screen "106_Rocno_postaja6" 1280x800, template "100_Rocno"
   IOField "I/O field_1" at 1132,158 size 125x32; FormatPattern 99999; Unit  l/min
      ProcessValue <- "FB_IOL_IFM_SV_DB_uPretok"
   IOField "I/O field_2" at 1132,210 size 128x32; FormatPattern 99.9; Unit  °C
      ProcessValue <- "FB_IOL_IFM_SV_DB_fTemperatura"
   TextField "Text field_2" at 1090,159 size 19x25; Text 'Q'
   TextField "Text field_3" at 1093,216 size 16x25; Text 'T'
   TextField "Text field_4" at 1144,120 size 58x25; Text 'VODA'
   IOField "I/O field_3" at 1132,304 size 125x32; FormatPattern 99.9; Unit  bar
      ProcessValue <- "FB_Lin_FESTO_PNEVMATIKA_PRITISK_Q_izhod"
   TextField "Text field_5" at 1090,305 size 17x25; Text 'P'
   TextField "Text field_7" at 1144,266 size 56x25; Text 'ZRAK'
   IOField "I/O field_4" at 1133,400 size 125x32; FormatPattern 99.9; Unit  bar
      ProcessValue <- "FB_FESTO_VPPM_DB_setstatZeljeniPritisk"
   TextField "Text field_6" at 1091,401 size 17x25; Text 'P'
   TextField "Text field_8" at 1100,360 size 169x25; Text 'P ZATISKOVANJA'
   TextField "Text field_17" at 613,544 size 239x46; Text 'POBIRANJE/NALAGANJE KOMADA'
   IOField "I/O field_7" at 742,605 size 133x35; FormatPattern 99.9; Unit  mm
      ProcessValue <- "DB_HMI_SDAT1_PozPobiranje"
   IOField "I/O field_8" at 739,666 size 136x35; FormatPattern 99.9; Unit  mm
      ProcessValue <- "DB_HMI_SDAT1_PozNalaganje"
   TextField "Text field_12" at 280,615 size 118x25; Text 'NALAGANJE'
   TextField "Text field_13" at 281,677 size 114x25; Text 'POBIRANJE'
   TextField "Text field_14" at 290,544 size 239x46; Text 'POBIRANJE/NALAGANJE PLOŠČICE'
   Circle "Circle_8" at 393,678 size 21x21
      Appearance <- "SDAT2_oPoz1Dosezena"
   Circle "Circle_7" at 394,618 size 21x21
      Appearance <- "SDAT2_oPoz2Dosezena"
   IOField "I/O field_10" at 421,670 size 136x32; FormatPattern 99.9; Unit  mm
      ProcessValue <- "DB_HMI_SDAT2_PozPobiranje"
   IOField "I/O field_9" at 425,613 size 133x32; FormatPattern 99.9; Unit  mm
      ProcessValue <- "DB_HMI_SDAT2_PozNalaganje"
   IOField "I/O field_12" at 422,709 size 136x32; FormatPattern 99.99; Unit  mm
      ProcessValue <- "SDAT2_out"
   TextField "Text field_11" at 434,112 size 84x25; Text 'Keyence'
   IOField "I/O field_13" at 432,190 size 109x32; FormatPattern 999999; Unit  mm
      ProcessValue <- "DB_KEYENCE_Elektroda_ZeljenaPozicija_POZ1"
   IOField "I/O field_14" at 432,244 size 109x32; FormatPattern 999999; Unit  mm
      ProcessValue <- "DB_KEYENCE_Elektroda_ZeljenaPozicija_POZ2"
   TextField "Text field_18" at 369,147 size 213x25; Text 'ELEKTRODA GOR/DOL'
   IOField "I/O field_17" at 432,290 size 109x32; FormatPattern 999999; Unit  mm
      ProcessValue <- "DB_KEYENCE_Elektroda_ZeljenaPozicija_POZ3_elektrodaStisnjena"
   IOField "I/O field_18" at 431,334 size 109x32; FormatPattern 999999; Unit  mm
      ProcessValue <- "DB_KEYENCE_Elektroda_ZeljenaPozicija_POZ4_elektrodaZavarjeno"
   TextField "Text field_9" at 282,194 size 81x25; Text 'ZGORAJ'
   TextField "Text field_19" at 282,339 size 117x25; Text 'ZAVARJENO'
   TextField "Text field_20" at 282,294 size 112x25; Text 'STISNJENO'
   TextField "Text field_21" at 282,248 size 99x25; Text 'HLAJENJE'
   Circle "Circle_1" at 398,195 size 20x20
      Appearance <- "FB_KEYENCE_GT2_ODMIKVARJENJA_oPoz1Dosezena"
   Circle "Circle_2" at 399,250 size 20x20
      Appearance <- "FB_KEYENCE_GT2_ODMIKVARJENJA_oPoz2Dosezena"
   Circle "Circle_3" at 401,296 size 20x20
      Appearance <- "FB_KEYENCE_GT2_ODMIKVARJENJA_oPoz3Dosezena"
   Circle "Circle_4" at 401,339 size 20x20
      Appearance <- "FB_KEYENCE_GT2_ODMIKVARJENJA_oPoz4Dosezena"
   IOField "I/O field_11" at 740,706 size 136x35; FormatPattern 99.99; Unit  mm
      ProcessValue <- "SDAT1_out"
   IOField "I/O field_6" at 531,408 size 128x32; FormatPattern 999999; Unit  mm
      ProcessValue <- "Keyence_OdmičniCilinderVarjenja"
   TextField "Text field_1" at 608,610 size 118x25; Text 'NALAGANJE'
   TextField "Text field_10" at 608,672 size 114x25; Text 'POBIRANJE'
   Circle "Circle_9" at 716,674 size 21x21
      Appearance <- "SDAT1_oPoz1Dosezena"
   Circle "Circle_10" at 719,612 size 21x21
      Appearance <- "SDAT1_oPoz2Dosezena"
   TextField "Text field_22" at 823,111 size 84x25; Text 'Keyence'
   TextField "Text field_23" at 691,147 size 268x25; Text 'ELEKTRODA NAZAJ/NAPREJ'
   TextField "Text field_24" at 687,194 size 67x25; Text 'NAZAJ'
   TextField "Text field_27" at 687,243 size 78x25; Text 'NAPREJ'
   IOField "I/O field_15" at 805,190 size 109x32; FormatPattern 999999; Unit  mm
      ProcessValue <- "DB_KEYENCE_Kroznik_ZeljenaPozicija_POZ1"
   IOField "I/O field_16" at 805,242 size 109x32; FormatPattern 999999; Unit  mm
      ProcessValue <- "DB_KEYENCE_Kroznik_ZeljenaPozicija_POZ2"
   IOField "I/O field_5" at 944,408 size 125x32; FormatPattern s999999; Unit  mm
      ProcessValue <- "Keyence_OdmičniCilinderKonusa"
   Circle "Circle_5" at 770,198 size 20x20
      Appearance <- "FB_KEYENCE_GT2_odmikKonusaKroznika_oPoz1Dosezena"
   Circle "Circle_6" at 770,245 size 20x20
      Appearance <- "FB_KEYENCE_GT2_odmikKonusaKroznika_oPoz2Dosezena"
   IOField "I/O field_19" at 564,190 size 105x32; FormatPattern 999999; Unit  mm
      ProcessValue <- "DB_KEYENCE_Elektroda_TOLERANCA{1}"
   IOField "I/O field_20" at 565,244 size 105x32; FormatPattern 999999; Unit  mm
      ProcessValue <- "DB_KEYENCE_Elektroda_TOLERANCA{2}"
   IOField "I/O field_21" at 564,290 size 105x32; FormatPattern 999999; Unit  mm
      ProcessValue <- "DB_KEYENCE_Elektroda_TOLERANCA{3}"
   IOField "I/O field_22" at 565,334 size 105x32; FormatPattern 999999; Unit  mm
      ProcessValue <- "DB_KEYENCE_Elektroda_TOLERANCA{4}"
   IOField "I/O field_23" at 954,190 size 106x32; FormatPattern 999999; Unit  mm
      ProcessValue <- "DB_KEYENCE_TOLERANCA{1}"
   IOField "I/O field_24" at 954,242 size 106x32; FormatPattern 999999; Unit  mm
      ProcessValue <- "DB_KEYENCE_TOLERANCA{2}"
   TextField "Text field_15" at 934,191 size 20x25; Text '+'
   TextField "Text field_16" at 937,205 size 13x25; Text '-'
   TextField "Text field_25" at 937,241 size 20x25; Text '+'
   TextField "Text field_26" at 940,255 size 13x25; Text '-'
   TextField "Text field_28" at 548,188 size 20x25; Text '+'
   TextField "Text field_29" at 551,202 size 13x25; Text '-'
   TextField "Text field_30" at 548,242 size 20x25; Text '+'
   TextField "Text field_31" at 551,256 size 13x25; Text '-'
   TextField "Text field_32" at 548,289 size 20x25; Text '+'
   TextField "Text field_33" at 551,303 size 13x25; Text '-'
   TextField "Text field_34" at 548,334 size 20x25; Text '+'
   TextField "Text field_35" at 551,348 size 13x25; Text '-'
   IOField "I/O field_25" at 1090,512 size 174x32; FormatPattern 99999; Unit  kos
      ProcessValue <- "DB_HMI_ČiščenjeElektrode_ZeljenoStevilo"
   TextField "Text field_36" at 1125,460 size 114x46; Text 'CISCENJE ELEKTRODE'

screen "41_Settings2" 1280x800, template "02_Settings"
   GraphicView "Graphic view_2" at 0,0 size 1280x800; Picture "PopUpBackground"
      Visibility <- "PopUpBackground"
   IOField "I/O field_1" at 1132,158 size 125x32; FormatPattern 99999; Unit  l/min
      ProcessValue <- "FB_IOL_IFM_SV_DB_uPretok"
   IOField "I/O field_2" at 1132,210 size 128x32; FormatPattern 99.9; Unit  °C
      ProcessValue <- "FB_IOL_IFM_SV_DB_fTemperatura"
   TextField "Text field_2" at 1090,159 size 19x25; Text 'Q'
   TextField "Text field_3" at 1093,216 size 16x25; Text 'T'
   TextField "Text field_4" at 1144,120 size 58x25; Text 'VODA'
   IOField "I/O field_3" at 1132,314 size 125x32; FormatPattern 99.9; Unit  bar
      ProcessValue <- "FB_Lin_FESTO_PNEVMATIKA_PRITISK_Q_izhod"
   TextField "Text field_5" at 1090,315 size 17x25; Text 'P'
   TextField "Text field_7" at 1144,276 size 56x25; Text 'ZRAK'
   IOField "I/O field_4" at 1132,470 size 125x32; FormatPattern 99.9; Unit  bar
      ProcessValue <- "FB_FESTO_VPPM_DB_setstatZeljeniPritisk"
   TextField "Text field_6" at 1090,471 size 17x25; Text 'P'
   TextField "Text field_8" at 1099,430 size 169x25; Text 'P ZATISKOVANJA'
   TextField "Text field_17" at 613,544 size 239x46; Text 'POBIRANJE/NALAGANJE KOMADA'
   Group "Group_2" at 606,112 size 282x342
   IOField "I/O field_7" at 742,605 size 133x35; FormatPattern 99.9; Unit  mm
      ProcessValue <- "DB_HMI_SDAT1_PozPobiranje"
   IOField "I/O field_8" at 739,666 size 136x35; FormatPattern 99.9; Unit  mm
      ProcessValue <- "DB_HMI_SDAT1_PozNalaganje"
   TextField "Text field_12" at 280,615 size 118x25; Text 'NALAGANJE'
   TextField "Text field_13" at 281,677 size 114x25; Text 'POBIRANJE'
   TextField "Text field_14" at 290,544 size 239x46; Text 'POBIRANJE/NALAGANJE PLOŠČICE'
   Circle "Circle_8" at 393,678 size 21x21
      Appearance <- "SDAT2_oPoz1Dosezena"
   Circle "Circle_7" at 394,618 size 21x21
      Appearance <- "SDAT2_oPoz2Dosezena"
   IOField "I/O field_10" at 421,670 size 136x32; FormatPattern 99.9; Unit  mm
      ProcessValue <- "DB_HMI_SDAT2_PozPobiranje"
   IOField "I/O field_9" at 425,613 size 133x32; FormatPattern 99.9; Unit  mm
      ProcessValue <- "DB_HMI_SDAT2_PozNalaganje"
   IOField "I/O field_12" at 422,709 size 136x32; FormatPattern 99.99; Unit  mm
      ProcessValue <- "SDAT2_out"
   TextField "Text field_11" at 387,114 size 84x25; Text 'Keyence'
   IOField "I/O field_13" at 432,190 size 125x32; FormatPattern 999999; Unit  um
      ProcessValue <- "DB_KEYENCE_Elektroda_ZeljenaPozicija_POZ1"
   IOField "I/O field_14" at 432,244 size 125x32; FormatPattern 999999; Unit  um
      ProcessValue <- "DB_KEYENCE_Elektroda_ZeljenaPozicija_POZ2"
   TextField "Text field_18" at 333,147 size 213x25; Text 'ELEKTRODA GOR/DOL'
   IOField "I/O field_17" at 432,290 size 125x32; FormatPattern 999999; Unit  um
      ProcessValue <- "DB_KEYENCE_Elektroda_ZeljenaPozicija_POZ3_elektrodaStisnjena"
   IOField "I/O field_18" at 431,334 size 125x32; FormatPattern 999999; Unit  um
      ProcessValue <- "DB_KEYENCE_Elektroda_ZeljenaPozicija_POZ4_elektrodaZavarjeno"
   TextField "Text field_9" at 318,194 size 81x25; Text 'ZGORAJ'
   TextField "Text field_19" at 282,339 size 117x25; Text 'ZAVARJENO'
   TextField "Text field_20" at 287,294 size 112x25; Text 'STISNJENO'
   TextField "Text field_21" at 300,248 size 99x25; Text 'HLAJENJE'
   Circle "Circle_1" at 398,195 size 20x20
      Appearance <- "FB_KEYENCE_GT2_ODMIKVARJENJA_oPoz1Dosezena"
   Circle "Circle_2" at 399,250 size 20x20
      Appearance <- "FB_KEYENCE_GT2_ODMIKVARJENJA_oPoz2Dosezena"
   Circle "Circle_3" at 401,296 size 20x20
      Appearance <- "FB_KEYENCE_GT2_ODMIKVARJENJA_oPoz3Dosezena"
   Circle "Circle_4" at 401,339 size 20x20
      Appearance <- "FB_KEYENCE_GT2_ODMIKVARJENJA_oPoz4Dosezena"
   IOField "I/O field_11" at 740,706 size 136x35; FormatPattern 99.99; Unit  mm
      ProcessValue <- "SDAT1_out"
   IOField "I/O field_6" at 428,406 size 128x32; FormatPattern s999999; Unit  um
      ProcessValue <- "Keyence_OdmičniCilinderVarjenja"
   TextField "Text field_1" at 608,610 size 118x25; Text 'NALAGANJE'
   TextField "Text field_10" at 608,672 size 114x25; Text 'POBIRANJE'
   Circle "Circle_9" at 716,674 size 21x21
      Appearance <- "SDAT1_oPoz1Dosezena"
   Circle "Circle_10" at 719,612 size 21x21
      Appearance <- "SDAT1_oPoz2Dosezena"
   TextField "Text field_22" at 703,114 size 84x25; Text 'Keyence'
   TextField "Text field_23" at 620,147 size 268x25; Text 'ELEKTRODA NAZAJ/NAPREJ'
   TextField "Text field_24" at 640,194 size 67x25; Text 'NAZAJ'
   TextField "Text field_27" at 635,243 size 78x25; Text 'NAPREJ'
   IOField "I/O field_15" at 748,190 size 125x32; FormatPattern 999999; Unit  um
      ProcessValue <- "DB_KEYENCE_Kroznik_ZeljenaPozicija_POZ1"
   IOField "I/O field_16" at 748,242 size 125x32; FormatPattern 999999; Unit  um
      ProcessValue <- "DB_KEYENCE_Kroznik_ZeljenaPozicija_POZ2"
   IOField "I/O field_5" at 748,405 size 125x32; FormatPattern s999999; Unit  um
      ProcessValue <- "Keyence_OdmičniCilinderKonusa"
   Circle "Circle_5" at 713,198 size 20x20
      Appearance <- "FB_KEYENCE_GT2_odmikKonusaKroznika_oPoz1Dosezena"
   Circle "Circle_6" at 713,245 size 20x20
      Appearance <- "FB_KEYENCE_GT2_odmikKonusaKroznika_oPoz2Dosezena"

PopupScreen "VARILNIK" 300x695
   Button "Button_1" at 48,52 size 188x72; TextOff 'RESET'
      on Release: ResetBit("DB_HMI_Varjenje_ResetWithWC")
      on Press: SetBit("DB_HMI_Varjenje_ResetWithWC")
   Button "Button_2" at 48,140 size 188x72; TextOff 'RESET + ZVAR'
   SymbolicIOField "Symbolic I/O field_1" at 43,271 size 201x29; TextOn '1'; TextOff '0'; TextList "BOSH"
      ProcessValue <- "StatusCode"
   TextField "Text field_1" at 51,99 size 176x23; Text 'Reset varilnika z WC'
   TextField "Text field_2" at 52,187 size 176x23; Text 'Reset varilnika z zvarom'
   TextField "Text field_3" at 43,244 size 176x23; Text 'STATUS VARILNIKA:'
   TextField "Text field_4" at 37,10 size 221x23; Text 'VARILNIK BOSH 6000'

PopupScreen "STEVCI" 810x660
   TextField "Text field_14" at 12,94 size 150x23; Text 'ŠTEVEC SKUPAJ'
   IOField "I/O field_5" at 193,93 size 133x32; FormatPattern 999999; Unit  KOS
      ProcessValue <- "DB_STEVCI_STEVCI_SKUPAJ"
   TextField "Text field_1" at 12,143 size 129x21; Text 'ZAVARJENO OK'
   TextField "Text field_2" at 12,182 size 141x21; Text 'ZAVARJENO NOK'
   IOField "I/O field_1" at 196,137 size 133x32; FormatPattern 999999; Unit  KOS
      ProcessValue <- "DB_STEVCI_STEVCI_ZavarjenoOK"
   IOField "I/O field_2" at 196,176 size 133x32; FormatPattern 999999; Unit  KOS
      ProcessValue <- "DB_STEVCI_STEVCI_ZavarjenoNOK"
   TextField "Text field_3" at 243,10 size 214x31; Text 'ŠTEVCI IZDELKOV'
   TextField "Text field_4" at 14,55 size 96x23; Text 'VARJENJE'
   TextField "Text field_5" at 404,94 size 150x23; Text 'ŠTEVEC SKUPAJ'
   IOField "I/O field_3" at 585,93 size 133x32; FormatPattern 999999; Unit  KOS
      ProcessValue <- "DB_STEVCI_STEVCI KAMERA_SKUPAJ"
   TextField "Text field_6" at 404,143 size 100x21; Text 'KAMERA OK'
   TextField "Text field_7" at 404,182 size 112x21; Text 'KAMERA NOK'
   IOField "I/O field_4" at 588,137 size 133x32; FormatPattern 999999; Unit  KOS
      ProcessValue <- "DB_STEVCI_STEVCI KAMERA_KameraOK"
   IOField "I/O field_6" at 588,176 size 133x32; FormatPattern 999999; Unit  KOS
      ProcessValue <- "DB_STEVCI_STEVCI KAMERA_KameraNOK"
   TextField "Text field_8" at 406,55 size 82x23; Text 'KAMERA'
   TextField "Text field_9" at 765,14 size 23x24; Text 'X'
   Button "btnPreviousScreen" at 744,0 size 66x55; TextOff 'Text'
      on Click: function_efd93a16("STEVCI", 0, 0, 0, -1, 1)

PopupScreen "RESETSKATEL" 300x695
   Button "Button_1_1" at 48,70 size 188x72; TextOff 'IZPRAZNI SKATLO 1'
      on Press: SetBit("DB_HMI_TekočiTrak_btnResetSkatle1")
      on Release: ResetBit("DB_HMI_TekočiTrak_btnResetSkatle1")
   Button "Button_2" at 43,279 size 188x72; TextOff 'IZPRAZNI SKATLO 2'
      on Press: SetBit("DB_HMI_TekočiTrak_btnResetSKatle2")
      on Release: ResetBit("DB_HMI_TekočiTrak_btnResetSKatle2")
   TextField "Text field_1" at 49,119 size 186x23; Text 'Reset stevca polne škatle'
   TextField "Text field_2" at 47,328 size 176x23; Text 'Reset števca polne škatle'
   TextField "Text field_3" at 16,154 size 176x23; Text 'STATUS :'
   TextField "Text field_4" at 10,10 size 281x23; Text 'SKATLA IZDELKOV POLNA'
   TextField "Text field_5" at 16,367 size 176x23; Text 'STATUS :'
   SymbolicIOField "Symbolic I/O field_1" at 79,155 size 191x22; TextOff '0'; TextOn '1'; TextList "StatusSkatel"
      ProcessValue <- "FB_TekociTrak_DB_stat_skatla1Polna"
   SymbolicIOField "Symbolic I/O field_2" at 79,368 size 191x22; TextOn '1'; TextOff '0'; TextList "StatusSkatel"
      ProcessValue <- "FB_TekociTrak_DB_stat_skatla2Polna"

VB script "ActivateAlarmControlScreen"
   bec8f1e5-2ab1-45f6-ad91-1d37c469eb91 20_Messages,0

VB script "ActivateStartScreen"
   HmiRuntime.BaseScreenName = SmartTags("StartScreenName")

VB script "CheckCurrentLanguage"
   If HmiRuntime.Language = 1031 Then 'German
   	SmartTags("CurrentLanguage") = 0
   	ElseIf HmiRuntime.Language = 1033 Then 'English US
   	SmartTags("CurrentLanguage") = 1
   End If
   
   	

VB script "CheckCurrentUserName"
   If SmartTags("CurrentUserName") = "" Or SmartTags("CurrentUserName") = "User Name" Or SmartTags("CurrentUserName") = "Benutzer" Then
     
     If HmiRuntime.Language = 1031 Then 'Germany
       SmartTags("CurrentUserName") = "Benutzer"
       
     ElseIf HmiRuntime.Language = 1033 Then 'English US
       SmartTags("CurrentUserName") = "User Name"
     End If
     
     SmartTags("UserIsLoggedIn") = False
   Else
     If SmartTags("CurrentUserName") <> "User Name" And SmartTags("CurrentUserName") <> "Benutzer" Then
       SmartTags("UserIsLoggedIn") = True  
     End If
   End If

VB script "CheckDiagState"
   If SmartTags("@DiagnosticsIndicatorTag") = 1 Then
   	SmartTags("DiagState") = 1
   Else
   	SmartTags("DiagState") = 0
   End If

VB script "GetStartScreenName"
   SmartTags("StartScreenName") = HmiRuntime.BaseScreenName

VB script "ShowLoginPopUp"
   efd93a16-2665-4b85-bcb9-25eddcb7b6f4 Template_Logon_Logoff,480,110,$3$hmiOn$,$3$hmiAnimationOff$,$3$hmiFast$

VB script "ShowOperatingModePopUp"
   efd93a16-2665-4b85-bcb9-25eddcb7b6f4 Template_Operating_Mode,428,110,$3$hmiOn$,$3$hmiAnimationOff$,$3$hmiFast$

VB script "ShowOptionPanelPopUp"
   efd93a16-2665-4b85-bcb9-25eddcb7b6f4 OptionPanel_4_Buttons, 890, 110, $3$hmiOn$, $3$hmiRight$, $3$hmiFast$

VB script "ShowRecipePopUp"
   efd93a16-2665-4b85-bcb9-25eddcb7b6f4 Template_Recipe,290,110,$3$hmiOn$,$3$hmiAnimationOff$,$3$hmiFast$

VB script "VBFunction_1"
   'Tip:
   ' 1. Use the <CTRL+SPACE> or <CTRL+I> shortcut to open a list of all objects and functions
   ' 2. Write the code using the HMI Runtime object.
   '  Example: HmiRuntime.Screens("Screen_1").
   ' 3. Use the <CTRL+J> shortcut to create an object reference.
   'Write the code as of this position:
   
   'Please replace all sequences which are enclosed with '_' by your own code.
   
   
   '1s trigger
   
   'Poglej ce je napaka Varjenja in prigaži meni
   
   'Rectangle_17
   
   'Dim btnResetSkatle1, btnResetSkatle2
   'Set btnResetSkatle1 = HmiRuntime.ActiveScreen.ScreenItems("Button_2")
   'Set btnResetSkatle2 = HmiRuntime.ActiveScreen.ScreenItems("Rectangle_17")
   'Set btnResetSkatle1 = HmiRuntime.Screens("Slide-in screen left").ScreenItems("Button_1")
   Dim activatescreen11
   Dim screenname,txt
   screenname = HmiRuntime.BaseScreenName
   
   'Set txt = HmiRuntime.ActiveScreen.ScreenItems("Text15")
   'txt.Text = screenname
   
   If  SmartTags("TimerReady") = 0  Then
   	'ShowSlideInScreen "Slide-in screen left", hmiOn
   	efd93a16-2665-4b85-bcb9-25eddcb7b6f4 VARILNIK,0,105,$3$hmiOn$,$3$hmiAnimationOff$,$3$hmiFast$
   	activatescreen11 = True
   	
   	
   Else
   	efd93a16-2665-4b85-bcb9-25eddcb7b6f4 VARILNIK,0,105,$3$hmiOff$,$3$hmiAnimationOff$,$3$hmiFast$
   	activatescreen11 = False
   End If
   
   
   
   'Please replace all sequences which are enclosed with '_' by your own code.
   If ((SmartTags("DB_STEVCI_STEVEC_SKATEL_SKATLA1") >= SmartTags("DB_STEVCI_STEVCI_ZELENAPOLNA_SKATLA_SKATLA1") Or (SmartTags("DB_STEVCI_STEVEC_SKATEL_SKATLA2") >= SmartTags("DB_STEVCI_STEVCI_ZELENAPOLNA_SKATLA_SKATLA2"))) And (Not activatescreen11)) Then
   	efd93a16-2665-4b85-bcb9-25eddcb7b6f4 RESETSKATEL,0,105,$3$hmiOn$,$3$hmiAnimationOff$,$3$hmiFast$
   	'btnResetSkatle1.Top = 10
   	'btnResetSkatle1.Visible = 1
   	'ModraSkatla
   	'btnResetSkatle2.BackColor = RGB(0,95,135)
   	
   	
   Else
   	efd93a16-2665-4b85-bcb9-25eddcb7b6f4 RESETSKATEL,0,105,$3$hmiOff$,$3$hmiAnimationOff$,$3$hmiFast$
   	'btnResetSkatle1.Visible = 0
   	'SivaSkatla
   	'btnResetSkatle2.BackColor = RGB(217, 217, 217)
   End If

VB script "VBFunction_2"
   'Tip:
   ' 1. Use the <CTRL+SPACE> or <CTRL+I> shortcut to open a list of all objects and functions
   ' 2. Write the code using the HMI Runtime object.
   '  Example: HmiRuntime.Screens("Screen_1").
   ' 3. Use the <CTRL+J> shortcut to create an object reference.
   'Write the code as of this position:

scheduled task "User Name"
   on Action: function_f41c6f6c("CurrentUserName"); "CheckCurrentUserName"()
*)